screen "praca" 800x480
   on GenerateScreen: SetTag("Tag_ScreenNumber", 5)
   GraphicView "Graphic view_4" at 274,396 size 70x70; Picture "soil-sensor_11298794"
   GraphicView "Graphic view_3" at 3,175 size 70x70; Picture "sensor_4212513"
   GraphicView "Graphic view_5" at 267,175 size 70x70; Picture "sensor_4212519"
   GraphicView "Graphic view_1" at 559,396 size 70x70; Picture "fan_4829316"
      Visibility <- "Wentylator"
   GraphicView "Graphic view_6" at 560,270 size 70x70; Picture "heater_4463010"
      Visibility <- "Grzałka"
   GraphicView "Graphic view_7" at 559,164 size 70x70; Picture "irrigation_18631825"
      Visibility <- "Pompa_podlewanie"
   GraphicView "Graphic view_8" at 11,397 size 70x70; Picture "anemometer_1113716"
   GraphicView "Graphic view_9" at 559,396 size 70x70; Picture "fan_off"
      Visibility <- "Wentylator"
   GraphicView "Graphic view_10" at 560,270 size 70x70; Picture "heater_off"
      Visibility <- "Grzałka"
   GraphicView "Graphic view_11" at 559,164 size 70x70; Picture "irrigation_off"
      Visibility <- "Pompa_podlewanie"
   GraphicView "Graphic view_12" at 278,267 size 70x70; Picture "sensor_2828470"
   TextField "Text field_1" at 52,152 size 204x23; Text 'INSOLATION / NASŁONECZNIENIE / SONNENEINSTRAHLUNG'
   TextField "Text field_3" at 44,373 size 166x23; Text 'SZYBKOŚĆ WIATRU'
   TextField "Text field_5" at 289,152 size 223x23; Text 'WILGOTNOŚĆ POWIETRZA'
   TextField "Text field_6" at 318,373 size 175x23; Text 'WILGOTNOŚĆ GLEBY'
   TextField "Text field_7" at 640,147 size 116x23; Text 'PODLEWANIE'
   TextField "Text field_8" at 635,256 size 80x23; Text 'GRZANIE'
   TextField "Text field_9" at 627,373 size 117x23; Text 'WENTYLACJA'
   TextField "Text field_10" at 81,3 size 256x34; Text 'PODGLĄD NA ŻYWO'
   Button "Button_1" at 750,0 size 50x50; TextOff 'WRÓĆ'; PictureOff "Back_arrow"
      on Click: function_efd93a16()
   Button "Button_2" at 3,1 size 43x43; TextOff 'DOM'; PictureOff "home_1"
      on Click: ActivateScreen("Root screen", 0)
   IOField "I/O field_3" at 94,402 size 70x65; FormatPattern 999
      ProcessValue <- "Czujnik_wiatru"
   IOField "I/O field_5" at 348,277 size 83x65; FormatPattern 9999
      ProcessValue <- "Zewnetrzny_czujnik_CO2"
   IOField "I/O field_4" at 377,172 size 69x65; FormatPattern 999
      ProcessValue <- "Czujnik_wilgotności_powietrza"
   IOField "I/O field_6" at 381,397 size 68x65; FormatPattern 999
      ProcessValue <- "Czujnik_wilgotności_gleby"
   TextField "Text field_12" at 446,190 size 47x46; Text '%'
   TextField "Text field_13" at 466,405 size 47x46; Text '%'
   TextField "Text field_14" at 192,164 size 47x72; Text 'W m²'
   IOField "I/O field_1" at 83,190 size 101x32; FormatPattern 99999
      ProcessValue <- "Czujnik_natezenia_światła"
   TextField "Text field_15" at 173,402 size 52x72; Text 'Km h'
   Circle "Circle_1" at 703,188 size 48x48
      Visibility <- "Pompa_podlewanie"
   Circle "Circle_2" at 702,283 size 48x48
      Visibility <- "Grzałka"
   TextField "Text field_16" at 447,283 size 69x39; Text 'ppm'
   Circle "Circle_4" at 703,188 size 48x48
      Visibility <- "Pompa_podlewanie"
   Circle "Circle_5" at 702,283 size 48x48
      Visibility <- "Grzałka"
   Circle "Circle_3" at 703,415 size 48x48
      Visibility <- "Wentylator"
   Circle "Circle_6" at 703,415 size 48x48
      Visibility <- "Wentylator"
   TextField "Text field_17" at 381,3 size 288x34; Text 'PODGLĄD NA ŻYWO / TRYB AUTOMATYCZNY'
      Visibility <- "HMI_Aktywacja_trybu_automatycznego"
   GraphicView "Graphic view_13" at 560,63 size 70x70; Picture "sprinkler_4552152"
      Visibility <- "Pompa_zraszacze"
   GraphicView "Graphic view_14" at 560,63 size 70x70; Picture "sprinkler"
      Visibility <- "Pompa_zraszacze"
   Circle "Circle_7" at 703,83 size 48x48
      Visibility <- "Pompa_zraszacze"
   Circle "Circle_8" at 703,83 size 48x48
      Visibility <- "Pompa_zraszacze"
   TextField "Text field_19" at 640,50 size 156x23; Text 'PODLEWANIE / MIKROZRASZANIE'
   GraphicView "Graphic view_15" at 0,66 size 70x70; Picture "Thermometer_icon"
   IOField "I/O field_8" at 73,73 size 97x65; FormatPattern 99.99
      ProcessValue <- "Temperatura_wewnetrzna"
   TextField "Text field_21" at 171,85 size 46x46; Text '°C'
   GraphicView "Graphic view_16" at 275,66 size 70x70; Picture "Thermometer_icon"
   IOField "I/O field_9" at 348,73 size 97x65; FormatPattern 99.99
      ProcessValue <- "Temperatura_zewnetrzna"
   TextField "Text field_23" at 447,82 size 46x46; Text '°C'
   TextField "Text field_20" at 57,44 size 137x42; Text 'TEMPERATURA TEMPERATURA WEWNTĘTRZNA'
   TextField "Text field_22" at 334,44 size 132x42; Text 'TEMPERATURA TEMPERATURA ZEWNĘTRZNA'
   GraphicView "Graphic view_2" at 11,273 size 70x70; Picture "sensor_2828470"
   IOField "I/O field_2" at 81,283 size 83x65; FormatPattern 9999
      ProcessValue <- "Wewnetrzny_czujnik_CO2"
   TextField "Text field_11" at 180,289 size 69x39; Text 'ppm'
   TextField "Text field_2" at 83,252 size 124x42; Text 'STĘŻENIE CO2 WEWNĘTRZNE STĘŻENIE CO2'
   TextField "Text field_4" at 352,256 size 123x42; Text 'STĘŻENIE CO2 ZEWNĘTRZNE STĘŻENIE CO2'
   TextField "Text field_18" at 381,3 size 211x34; Text 'TRYB RECEPTUR'
      Visibility <- "HMI_Aktywacja_trybu_Receptur"

Template "Template_1" 800x480
   Button "Exit" at 671,429 size 71x50; TextOn 'Exit'; TextOff 'Exit'; PictureOn "ExitRuntime_KTP700_Basic_PN_TR"; PictureOff "ExitRuntime_KTP700_Basic_PN_TR"
      on Release: StopRuntime(0)
   Button "Alarms" at 524,429 size 71x50; TextOn 'Alarms'; TextOff 'Alarms'; PictureOn "AlarmDisplay_KTP700_Basic_PN_TR"; PictureOff "AlarmDisplay_KTP700_Basic_PN_TR"
      on Release: function_ef3f5d25("Alarm window_Unacknowledged", -1)
   Button "Start screen" at 169,429 size 71x50; TextOn 'Start screen'; TextOff 'Start screen'; PictureOn "NavigateHome_KTP700_Basic_PN_TR"; PictureOff "NavigateHome_KTP700_Basic_PN_TR"
      on Release: ActivateScreen("Root screen", 0)
      Visibility <- "AlwaysTRUE"
   Button "Language" at 377,429 size 71x50; TextOn 'Language'; TextOff 'Language'; PictureOn "ToggleLanguage_KTP700_Basic_PN_TR"; PictureOff "ToggleLanguage_KTP700_Basic_PN_TR"
      on Release: function_fb9197e8(-1)

screen "Receptury" 800x480
   RecipeView "Recipe view_1" at 0,38 size 799x413; Recipe "Receptura_nr1"; RecipeNameCaption 'Recipe Name: / Wybierz Recepturę / Rezepturname:'; EntryNameCaption 'Entry Name / Zapisane Parametry / Eintragsname'; DataRecordNameCaption 'Data Record Name: / Wybierz Recepturę / Datensatzname:'
   GraphicView "Graphic view_1" at 529,152 size 35x35; Picture "Thermometer_icon"
   GraphicView "Graphic view_2" at 529,190 size 35x35; Picture "sensor_4212519"
   GraphicView "Graphic view_3" at 529,230 size 35x35; Picture "soil-sensor_11298794"
   GraphicView "Graphic view_4" at 529,269 size 35x35; Picture "window_11250237"
   GraphicView "Graphic view_5" at 529,308 size 35x35; Picture "sensor_2828470"
   GraphicView "Graphic view_6" at 529,348 size 35x35; Picture "sensor_4212513"
   TextField "Text field_11" at 569,150 size 39x38; Text '°C'
   TextField "Text field_18" at 569,190 size 39x38; Text '%'
   TextField "Text field_1" at 569,230 size 39x38; Text '%'
   TextField "Text field_2" at 564,269 size 57x32; Text '1/0'
   TextField "Text field_16" at 563,308 size 55x32; Text 'ppm'
   TextField "Text field_6" at 576,339 size 28x50; Text '°C W m'
   TextField "Text field_3" at 593,362 size 31x17; Text '2'
   Button "Button_1" at 750,0 size 50x50; TextOff 'WRÓĆ'; PictureOff "Back_arrow"
      on Click: function_efd93a16()
   Button "Button_14" at 3,1 size 43x43; TextOff 'DOM'; PictureOff "home_1"
      on Click: ActivateScreen("Root screen", 0)
   TextField "Text field_4" at 320,2 size 170x37; Text 'RECEPTURY'
   TextField "Text field_5" at 12,448 size 50x23; Text 'Nowy'
   TextField "Text field_7" at 69,448 size 57x23; Text 'Zapisz'
   TextField "Text field_8" at 137,448 size 45x23; Text 'Usuń'
   TextField "Text field_9" at 190,438 size 60x42; Text 'Zmień Nazwę'
   TextField "Text field_10" at 663,438 size 66x42; Text 'Załaduj z PLC'
   TextField "Text field_12" at 729,438 size 66x42; Text 'Załaduj do PLC'
   Button "Button_2" at 405,402 size 255x40; TextOff 'ZATWIERDŹ'
      on Click: ActivateScreen("praca", 0)
   TextField "Text field_13" at 456,450 size 173x23; Text 'Przejdź w tryb pracy'
   Button "Button_3" at 256,401 size 140x40; TextOff 'Z'
      on Click: function_ea909784(1, U 0, '\USB_X60.1\record.csv', 2, 1, N)
   TextField "Text field_14" at 266,438 size 113x42; Text 'Zapisz Kopię zapasową'

screen "Symulacja_czujnikow" 800x480
   TextField "Text field_1" at 21,47 size 252x23; Text 'Czujnik Wilgotności powietrza'
   TextField "Text field_2" at 308,47 size 214x23; Text 'Czujnik Wilgotności gleby'
   TextField "Text field_3" at 32,202 size 202x23; Text 'Termometr wewnętrzny'
   TextField "Text field_4" at 323,202 size 197x23; Text 'Termometr zewnętrzny'
   TextField "Text field_5" at 569,47 size 216x23; Text 'Czujnik natężenia światła'
   TextField "Text field_6" at 607,202 size 124x23; Text 'Czujnik wiatru'
   TextField "Text field_7" at 27,346 size 208x23; Text 'Wewnętrzny czujnik CO2'
   TextField "Text field_8" at 306,346 size 202x23; Text 'Zewnętrzny czujnik CO2'
   TextField "Text field_9" at 569,346 size 206x23; Text 'Stopień zasłonięcia rolet'
   IOField "I/O field_4" at 599,83 size 150x60; FormatPattern 9999
      ProcessValue <- "Czujnik_natezenia_światła"
   IOField "I/O field_5" at 599,242 size 150x60; FormatPattern 999
      ProcessValue <- "Czujnik_wiatru"
   IOField "I/O field_6" at 69,375 size 150x60; FormatPattern 9999
      ProcessValue <- "Wewnetrzny_czujnik_CO2"
   IOField "I/O field_7" at 346,375 size 150x60; FormatPattern 9999
      ProcessValue <- "Zewnetrzny_czujnik_CO2"
   IOField "I/O field_8" at 599,375 size 150x60; FormatPattern 999
      ProcessValue <- "Stopien_zasloniecia_rolet"
   IOField "I/O field_10" at 69,83 size 150x60; FormatPattern 999
      ProcessValue <- "Czujnik_wilgotności_powietrza"
   IOField "I/O field_11" at 346,83 size 150x60; FormatPattern 999
      ProcessValue <- "Czujnik_wilgotności_gleby"
   IOField "I/O field_12" at 69,242 size 150x60; FormatPattern 99.9
      ProcessValue <- "Temperatura_wewnetrzna"
   IOField "I/O field_13" at 346,242 size 150x60; FormatPattern 99.9
      ProcessValue <- "Temperatura_zewnetrzna"
   TextField "Text field_10" at 248,5 size 321x34; Text 'ZAPISZ RECEPTURE / SYMULACJA CZUJNIKÓW'
   Button "Button_1" at 750,0 size 50x50; TextOff 'WRÓĆ'; PictureOff "Back_arrow"
      on Click: function_efd93a16()
   Button "Button_14" at 3,1 size 43x43; TextOff 'DOM'; PictureOff "home_1"
      on Click: ActivateScreen("Root screen", 0)

screen "tryb_automatyczny" 800x480
   on GenerateScreen: SetTag("Tag_ScreenNumber", 1)
   IOField "I/O field_1" at 100,354 size 57x40; FormatPattern 99.9
      ProcessValue <- "Temperatura_wewnetrzna"
   Button "Button_1" at 750,0 size 50x50; TextOff 'WRÓĆ'; PictureOff "Back_arrow"
      on Click: function_efd93a16()
   Button "Button_2" at 504,411 size 285x60; TextOff 'ZATWIERDŹ'
      on Click: SetBit("HMI_Aktywacja_trybu_automatycznego"); ActivateScreen("praca", 0)
   Bar "Bar_1" at 14,103 size 70x275; MinimumValue 0; MaximumValue 45
      ProcessValue <- "Temperatura_auto"
   TextField "Text field_2" at 15,60 size 132x23; Text 'TEMPERATURA'
   Bar "Bar_2" at 217,108 size 70x275; MinimumValue 0; MaximumValue 100
      ProcessValue <- "Wilgotnosc_powietrza_auto"
   TextField "Text field_3" at 205,61 size 122x42; Text 'WOLGOTNOŚĆ POWIETRZA WILGOTNOŚĆ POWIETRZA'
   Button "Button_3" at 90,119 size 75x45; TextOff '+ / +0.5 °C'
      on Press: function_dd21b452("Temperatura_auto", 0.5)
   Button "Button_7" at 89,177 size 75x45; TextOff '- / -0.5 °C'
      on Press: function_b9b71300("Temperatura_auto", 0.5)
   IOField "I/O field_2" at 100,276 size 62x40; FormatPattern 99.9
      ProcessValue <- "Temperatura_auto"
   TextField "Text field_11" at 155,285 size 23x22; Text '°C'
   TextField "Text field_9" at 155,358 size 23x22; Text '°C'
   Bar "Bar_4" at 417,105 size 70x275; MinimumValue 0; MaximumValue 100
      ProcessValue <- "Wilgotnosc_gleby_auto"
   TextField "Text field_10" at 404,58 size 122x42; Text 'WOLGOTNOŚĆ GLEBY WILGOTNOŚĆ GLEBY'
   Button "Button_8" at 496,125 size 65x40; TextOff '+ / +2%'
      on Click: function_dd21b452("Wilgotnosc_gleby_auto", 2)
   Button "Button_9" at 497,177 size 65x40; TextOff '- / -2%'
      on Click: function_b9b71300("Wilgotnosc_gleby_auto", 2)
   IOField "I/O field_5" at 510,276 size 60x40; FormatPattern 999
      ProcessValue <- "Wilgotnosc_gleby_auto"
   IOField "I/O field_6" at 512,346 size 58x40; FormatPattern 999
      ProcessValue <- "Czujnik_wilgotności_gleby"
   TextField "Text field_12" at 493,264 size 101x22; Text 'USTAWIONA'
   TextField "Text field_13" at 497,335 size 86x22; Text 'AKTUALNA'
   TextField "Text field_14" at 547,285 size 23x22; Text '%'
   TextField "Text field_15" at 547,356 size 23x22; Text '%'
   Button "Button_10" at 298,125 size 65x40; TextOff '+ / +5%'
      on Click: function_dd21b452("Wilgotnosc_powietrza_auto", 5)
   Button "Button_11" at 298,177 size 65x40; TextOff '- / -5%'
      on Click: function_b9b71300("Wilgotnosc_powietrza_auto", 5)
   IOField "I/O field_4" at 305,277 size 66x40; FormatPattern 999
      ProcessValue <- "Wilgotnosc_powietrza_auto"
   IOField "I/O field_7" at 307,349 size 62x40; FormatPattern 999
      ProcessValue <- "Czujnik_wilgotności_powietrza"
   TextField "Text field_16" at 292,264 size 101x22; Text 'USTAWIONA'
   TextField "Text field_17" at 294,335 size 86x22; Text 'AKTUALNA'
   TextField "Text field_18" at 346,286 size 23x22; Text '%'
   TextField "Text field_19" at 346,357 size 23x22; Text '%'
   Button "Button_14" at 3,1 size 43x43; TextOff 'DOM'; PictureOff "home_1"
      on Click: ActivateScreen("Root screen", 0)
   TextField "Text field_4" at 0,403 size 128x23; Text 'SYSTEM OKIEN'
   Switch "Switch_1" at 23,433 size 70x38; TextOn 'ON'; CaptionText 'Switch'; TextOff 'OFF'
      ProcessValue <- "System_okien_auto"
   GraphicView "Graphic view_1" at 150,60 size 40x40; Picture "Thermometer_icon"
   GraphicView "Graphic view_2" at 330,61 size 40x40; Picture "sensor_4212519"
   TextField "Text field_5" at 93,334 size 86x22; Text 'AKTUALNA'
   TextField "Text field_6" at 90,262 size 101x22; Text 'USTAWIONA'
   GraphicView "Graphic view_3" at 526,61 size 40x40; Picture "soil-sensor_11298794"
   TextField "Text field_1" at 250,4 size 288x34; Text 'TRYB AUTOMATYCZNY'
   Bar "Bar_3" at 620,105 size 70x275; MinimumValue 0; MaximumValue 1500
      ProcessValue <- "Naslonecznienie_auto"
   TextField "Text field_7" at 604,53 size 161x42; Text 'WOLGOTNOŚĆ GLEBY NASŁONECZNIENIE'
   GraphicView "Graphic view_4" at 725,79 size 40x40; Picture "sensor_4212513"
   Button "Button_4" at 696,125 size 65x40; TextOff '+ +50 W m'
      on Click: function_dd21b452("Naslonecznienie_auto", 50)
   Button "Button_5" at 697,177 size 65x40; TextOff '- -50 W m'
      on Click: function_b9b71300("Naslonecznienie_auto", 50)
   IOField "I/O field_3" at 709,276 size 61x40; FormatPattern 9999
      ProcessValue <- "Naslonecznienie_auto"
   TextField "Text field_8" at 693,264 size 101x22; Text 'USTAWIONA / USTAWIONE'
   IOField "I/O field_8" at 711,347 size 62x40; FormatPattern 9999
      ProcessValue <- "Czujnik_natezenia_światła"
   TextField "Text field_20" at 697,335 size 86x22; Text 'AKTUALNA / AKTUALNE'
   TextField "Text field_23" at 751,143 size 32x18; Text '2'
   TextField "Text field_24" at 748,196 size 32x18; Text '2'
   Bar "Bar_5" at 165,432 size 223x39; MinimumValue 400; MaximumValue 950
      ProcessValue <- "Poziom_CO2_auto"
   TextField "Text field_21" at 238,402 size 128x23; Text 'SYSTEM OKIEN / POZIOM CO2'
   IOField "I/O field_9" at 416,402 size 66x40; FormatPattern 999
      ProcessValue <- "Poziom_CO2_auto"
   TextField "Text field_22" at 386,394 size 101x22; Text 'USTAWIONA'
   IOField "I/O field_10" at 404,440 size 62x40; FormatPattern 999
      ProcessValue <- "Wewnetrzny_czujnik_CO2"
   TextField "Text field_25" at 397,425 size 86x22; Text 'AKTUALNA'
   Button "Button_6" at 155,400 size 65x40; TextOff '+ / +25ppm'
      on Click: function_dd21b452("Poziom_CO2_auto", 25)
   Button "Button_12" at 132,431 size 65x40; TextOff '+ / -25ppm'
      on Click: function_b9b71300("Poziom_CO2_auto", 25)
*)